(* Logix 5000 project; controller _GigaDiscovery vendor 1 type 14 code 244 rev 35.11; software revision 35.03 *) (continued)
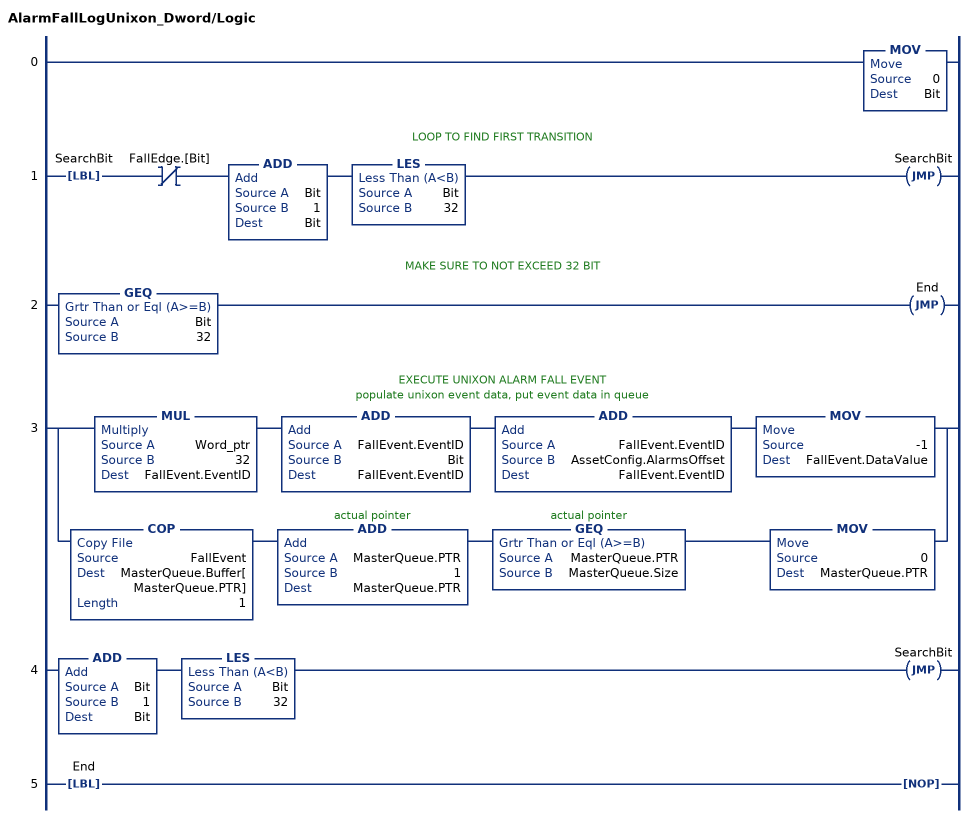
   0: MOV(0,Bit);
   // LOOP TO FIND FIRST TRANSITION
   1: LBL(SearchBit)XIO(FallEdge.[Bit])ADD(Bit,1,Bit)LES(Bit,32)JMP(SearchBit);
   // MAKE SURE TO NOT EXCEED 32 BIT
   2: GEQ(Bit,32)JMP(End);
   // EXECUTE UNIXON ALARM FALL EVENT
   // populate unixon event data, put event data in queue
   3: [MUL(Word_ptr,32,FallEvent.EventID) ADD(FallEvent.EventID,Bit,FallEvent.EventID) ADD(FallEvent.EventID,AssetConfig.AlarmsOffset,FallEvent.EventID) MOV(-1,FallEvent.DataValue) ,COP(FallEvent,MasterQueue.Buffer[MasterQueue.PTR],1) ADD(MasterQueue.PTR,1,MasterQueue.PTR) GEQ(MasterQueue.PTR,MasterQueue.Size) MOV(0,MasterQueue.PTR) ];
   4: ADD(Bit,1,Bit)LES(Bit,32)JMP(SearchBit);
   5: LBL(End)NOP();
END_ROUTINE
END_ADD_ON_INSTRUCTION

ADD_ON_INSTRUCTION AOI_DCM   (* revision 1.0 *)
VAR_INPUT
   Input_Type : BOOL; {required}   // 0 = Equivalent 1 = Complementary
   Discrepancy_Time : DINT; {required}   // (Msec)
   Channel_A : BOOL; {required}
   Channel_B : BOOL; {required}
   Channel_A_Status : BOOL; {required}
   Channel_B_Status : BOOL; {required}
   Reset_Pulse : BOOL; {required}
END_VAR
VAR_OUTPUT
   O1 : BOOL; {access Read Only, visible}
   FP : BOOL; {visible}
END_VAR
VAR
   Discrepancy_Timer : TIMER; {access None}
   Os : BOOL; {access None}
END_VAR

ROUTINE Logic   (* ladder *)
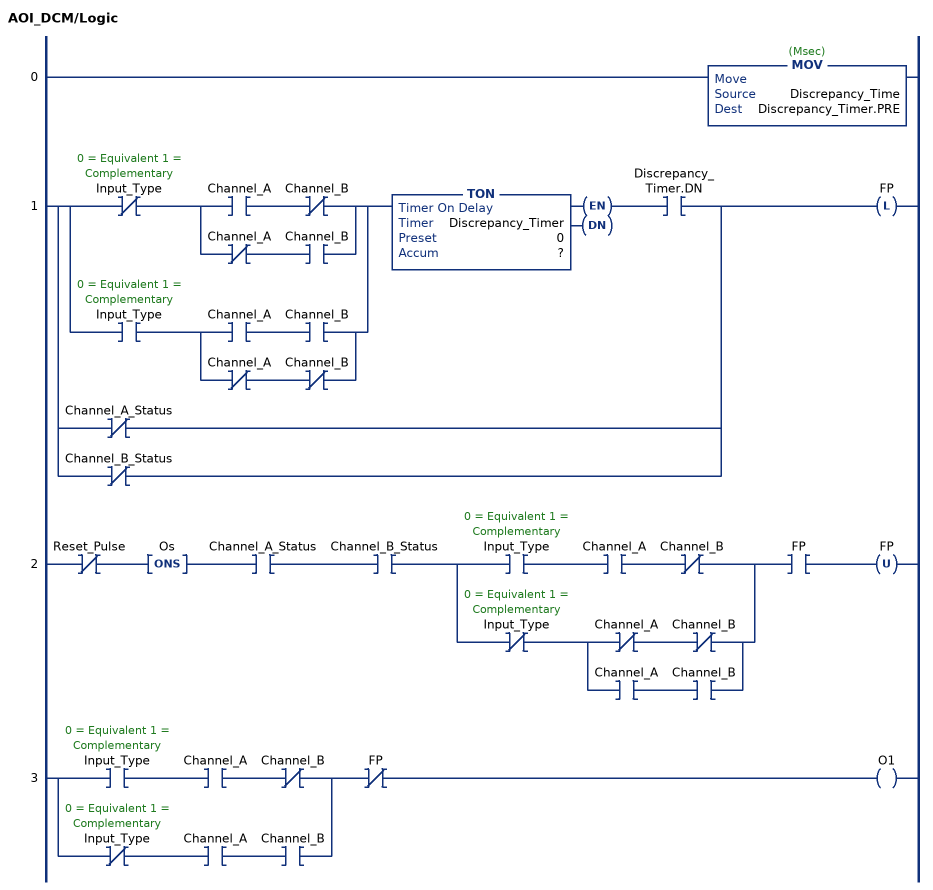
   0: MOV(Discrepancy_Time,Discrepancy_Timer.PRE);
   1: [[XIO(Input_Type) [XIC(Channel_A) XIO(Channel_B) ,XIO(Channel_A) XIC(Channel_B) ] ,XIC(Input_Type) [XIC(Channel_A) XIC(Channel_B) ,XIO(Channel_A) XIO(Channel_B) ] ] TON(Discrepancy_Timer,?,?) XIC(Discrepancy_Timer.DN) ,XIO(Channel_A_Status) ,XIO(Channel_B_Status) ]OTL(FP);
   2: XIO(Reset_Pulse)ONS(Os)XIC(Channel_A_Status)XIC(Channel_B_Status)[XIC(Input_Type) XIC(Channel_A) XIO(Channel_B) ,XIO(Input_Type) [XIO(Channel_A) XIO(Channel_B) ,XIC(Channel_A) XIC(Channel_B) ] ]XIC(FP)OTU(FP);
   3: [XIC(Input_Type) XIC(Channel_A) XIO(Channel_B) ,XIO(Input_Type) XIC(Channel_A) XIC(Channel_B) ]XIO(FP)OTE(O1);
END_ROUTINE
END_ADD_ON_INSTRUCTION

ADD_ON_INSTRUCTION EStop_AOI   (* revision 1.0, vendor Auxel *)
// Test the E-Stop Push Botton
// Revision note:
// Preliminary
// Help:
// This AOI request at the operator to check hte E-Stop function in cold mode (Ride not in start mode)
VAR_INPUT
   InEStopPbCh1 : BOOL; {access None, required}
   InEStopPbCh2 : BOOL; {required}
   InStatusCh1 : BOOL; {required}
   InStatusCh2 : BOOL; {required}
   cmdFltRst : BOOL; {required}
END_VAR
VAR_OUTPUT
   Test_Ok : BOOL; {access Read Only, visible}   // Test succefuly
   O1 : BOOL; {visible}
   FP : BOOL; {access Read Only, visible}
END_VAR
VAR
   Os : DINT; {access None}
   Sequencer : DINT; {access None}
   DCIS : DCI_STOP; {access None}
   In_Status : BOOL; {access None}
   PowerON : TIMER := (PRE := 200); {access None}
END_VAR

ROUTINE Logic   (* ladder *)
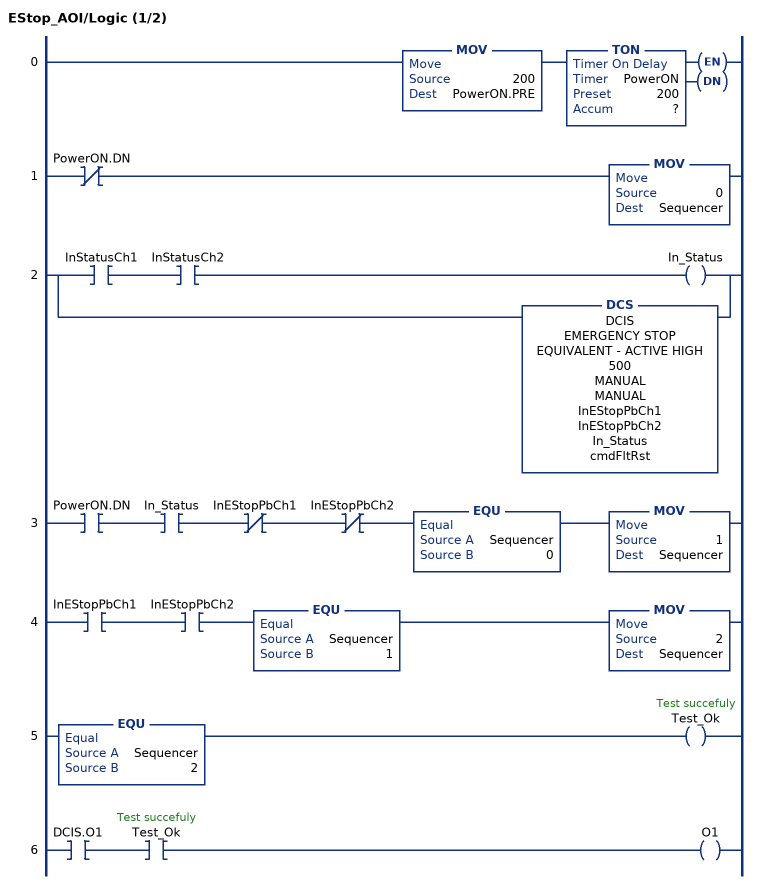
   0: MOV(200,PowerON.PRE)TON(PowerON,?,?);
   1: XIO(PowerON.DN)MOV(0,Sequencer);
   2: [XIC(InStatusCh1) XIC(InStatusCh2) OTE(In_Status) ,DCS(DCIS,EMERGENCY STOP,EQUIVALENT - ACTIVE HIGH,500,MANUAL,MANUAL,InEStopPbCh1,InEStopPbCh2,In_Status,cmdFltRst) ];
   3: XIC(PowerON.DN)XIC(In_Status)XIO(InEStopPbCh1)XIO(InEStopPbCh2)EQU(Sequencer,0)MOV(1,Sequencer);
   4: XIC(InEStopPbCh1)XIC(InEStopPbCh2)EQU(Sequencer,1)MOV(2,Sequencer);
   5: EQU(Sequencer,2)OTE(Test_Ok);
   6: XIC(DCIS.O1)XIC(Test_Ok)OTE(O1);
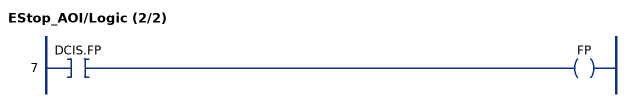
   7: XIC(DCIS.FP)OTE(FP);
END_ROUTINE
END_ADD_ON_INSTRUCTION

ADD_ON_INSTRUCTION Life_of_Machine   (* revision 1.0 *)
VAR_INPUT
   Start_Stop_Cycle_Started : BOOL; {required}
   HMI_Reset_Partial_Life_RunHH : BOOL; {required}
   HMI_Reset_Partial_Life_Cycle : BOOL; {required}
END_VAR
VAR_OUTPUT
   Life_HH : DINT; {access Read Only, visible}
   Partial_Life_HH : DINT; {access Read Only, visible}
   Working_Cycle_Number_Partial : DINT; {access Read Only, visible}
   Working_Cycle_Number_Total : DINT; {access Read Only, visible}
   Working_HH_Partial : DINT; {access Read Only, visible}
   Working_HH_Total : DINT; {access Read Only, visible}
   Working_Minutes_Partial : DINT; {access Read Only, visible}
END_VAR
VAR_INPUT
   HMI_Reset_Life_of_Machine : BOOL;
END_VAR
VAR
   Life_Hours : TIMER := (PRE := 3600000, ACC := 2467243); {access None}
   Life_HH_CTU : COUNTER; {access None}
   Partial_Life_HH_CTU : COUNTER; {access None}
   Working_Hours : TIMER := (PRE := 3600000, ACC := 2768993); {access None}
   Working_Minutes : TIMER := (PRE := 60000, ACC := 4300); {access None}
   Working_Cycle_Number_Partial_CTU : COUNTER; {access None}
   Working_Cycle_Number_Total_CTU : COUNTER; {access None}
   Working_HH_Partial_CTU : COUNTER; {access None}
   Working_HH_Total_CTU : COUNTER; {access None}
   Working_Minutes_Partial_CTU : COUNTER; {access None}
   Os : DINT; {access None}
END_VAR

ROUTINE Logic   (* ladder *)
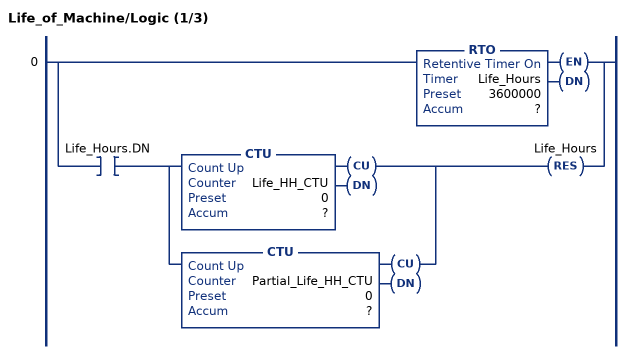
   0: [RTO(Life_Hours,?,?) ,XIC(Life_Hours.DN) [CTU(Life_HH_CTU,?,?) ,CTU(Partial_Life_HH_CTU,?,?) ] RES(Life_Hours) ];
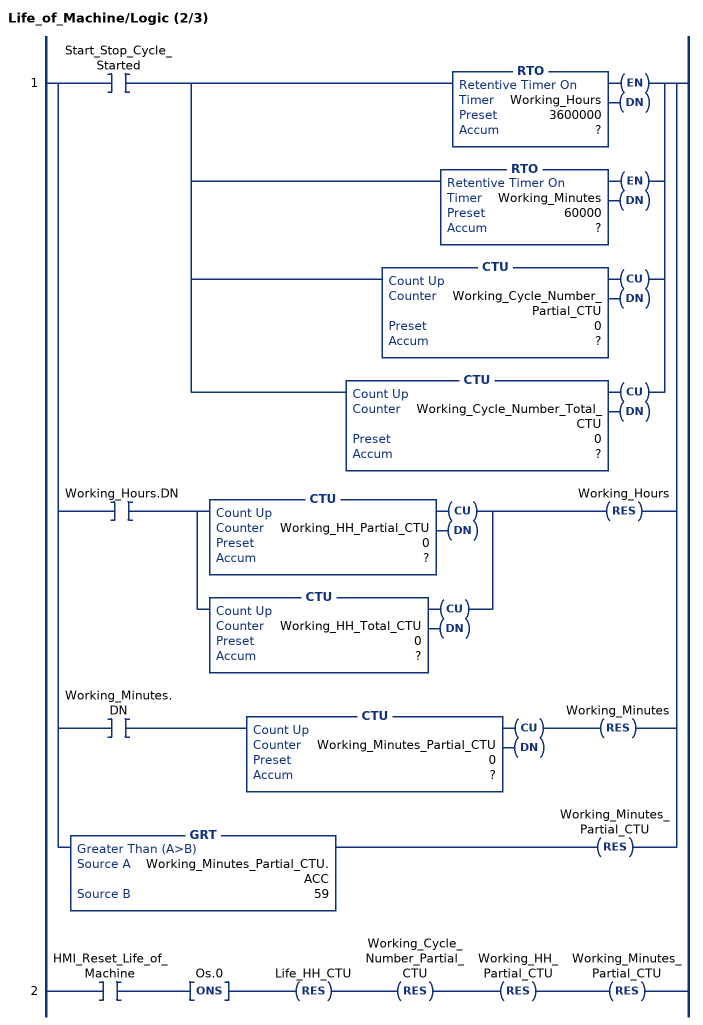
   1: [XIC(Start_Stop_Cycle_Started) [RTO(Working_Hours,?,?) ,RTO(Working_Minutes,?,?) ,[CTU(Working_Cycle_Number_Partial_CTU,?,?) ,CTU(Working_Cycle_Number_Total_CTU,?,?) ] ] ,XIC(Working_Hours.DN) [CTU(Working_HH_Partial_CTU,?,?) ,CTU(Working_HH_Total_CTU,?,?) ] RES(Working_Hours) ,XIC(Working_Minutes.DN) CTU(Working_Minutes_Partial_CTU,?,?) RES(Working_Minutes) ,GRT(Working_Minutes_Partial_CTU.ACC,59) RES(Working_Minutes_Partial_CTU) ];
   2: XIC(HMI_Reset_Life_of_Machine)ONS(Os.0)RES(Life_HH_CTU)RES(Working_Cycle_Number_Partial_CTU)RES(Working_HH_Partial_CTU)RES(Working_Minutes_Partial_CTU);
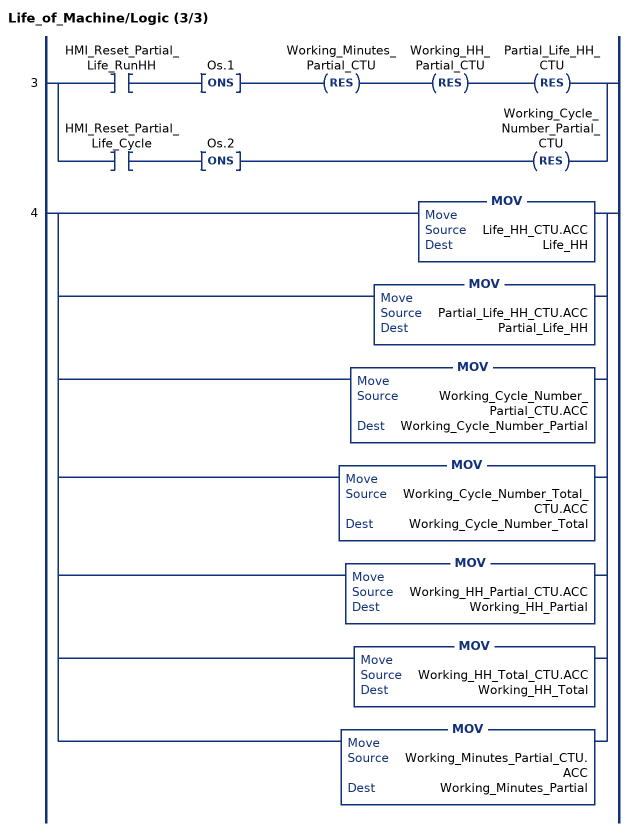
   3: [XIC(HMI_Reset_Partial_Life_RunHH) ONS(Os.1) RES(Working_Minutes_Partial_CTU) RES(Working_HH_Partial_CTU) RES(Partial_Life_HH_CTU) ,XIC(HMI_Reset_Partial_Life_Cycle) ONS(Os.2) RES(Working_Cycle_Number_Partial_CTU) ];
   4: [MOV(Life_HH_CTU.ACC,Life_HH) ,MOV(Partial_Life_HH_CTU.ACC,Partial_Life_HH) ,MOV(Working_Cycle_Number_Partial_CTU.ACC,Working_Cycle_Number_Partial) ,MOV(Working_Cycle_Number_Total_CTU.ACC,Working_Cycle_Number_Total) ,MOV(Working_HH_Partial_CTU.ACC,Working_HH_Partial) ,MOV(Working_HH_Total_CTU.ACC,Working_HH_Total) ,MOV(Working_Minutes_Partial_CTU.ACC,Working_Minutes_Partial) ];
END_ROUTINE
END_ADD_ON_INSTRUCTION

ADD_ON_INSTRUCTION Powerflex_DC_Fault   (* revision 1.0 *)
VAR_INPUT
   Fault_Code : DINT; {required}
END_VAR
VAR_IN_OUT
   Fault_Descrpition : STRING; {required}
END_VAR
VAR
   Fault_Descrpition_4 : STRING := 'AC Undervoltage'; {access None}
   Fault_Descrpition_5 : STRING := 'Arm Overvoltage'; {access None}
   Fault_Descrpition_2 : STRING := 'Auxiliary Input'; {access None}
   Fault_Descrpition_64 : STRING := 'Drive Overload'; {access None}
   Fault_Descrpition_132 : STRING := 'Dsp Error'; {access None}
   Fault_Descrpition_100 : STRING := '100'; {access None}
   Fault_Descrpition_32 : STRING; {access None}
   Fault_Descrpition_6 : STRING := 'Fld Current Loss'; {access None}
   Fault_Descrpition_95 : STRING := 'Fwd End Limit'; {access None}
   Fault_Descrpition_97 : STRING := 'Fwd Over Travel'; {access None}
   Fault_Descrpition_130 : STRING := 'Hardware Fault'; {access None}
   Fault_Descrpition_131 : STRING := 'Interrupt Error'; {access None}
   Fault_Descrpition_37 : STRING := 'Inverting Fault'; {access None}
   Fault_Descrpition_10 : STRING := 'Main Contactor'; {access None}
   Fault_Descrpition_7 : STRING := 'Motor Overload'; {access None}
   Fault_Descrpition_16 : STRING := 'Motor Over Temp'; {access None}
   Fault_Descrpition_90 : STRING := 'Open SCR'; {access None}
   Fault_Descrpition_13 : STRING := 'Overcurrent'; {access None}
   Fault_Descrpition_25 : STRING := 'Overspeed'; {access None}
   Fault_Descrpition_48 : STRING := 'Params Defaulted'; {access None}
   Fault_Descrpition_71 : STRING := 'Pommunication card fault Port 1'; {access None}
   Fault_Descrpition_81 : STRING := 'DPI port 1 stopped communicating'; {access None}
   Fault_Descrpition_93 : STRING := 'Resolver Error'; {access None}
   Fault_Descrpition_96 : STRING := 'Rev End Limit'; {access None}
   Fault_Descrpition_98 : STRING := 'Rev Over Travel'; {access None}
   Fault_Descrpition_89 : STRING := 'Shorted SCR'; {access None}
   Fault_Descrpition_91 : STRING := 'Spd Fdbk Loss'; {access None}
   Fault_Descrpition_62 : STRING := 'STune Aborted'; {access None}
   Fault_Descrpition_59 : STRING := 'STune CurLimit'; {access None}
   Fault_Descrpition_60 : STRING := 'STune FrictionLo'; {access None}
   Fault_Descrpition_58 : STRING := 'STune LoadHi'; {access None}
   Fault_Descrpition_56 : STRING := 'STune Overspeed'; {access None}
   Fault_Descrpition_57 : STRING := 'STune Stalled'; {access None}
   Fault_Descrpition_61 : STRING := 'STune Timeout'; {access None}
   Fault_Descrpition_70 : STRING := 'Sustained Curr'; {access None}
   Fault_Descrpition_94 : STRING := 'TorqPrv Spd Band'; {access None}
   Fault_Descrpition_99 : STRING := 'Travel Lim Cflct'; {access None}
   Fault_Descrpition_92 : STRING := 'Encoder Error'; {access None}
   Fault_Descrpition_8 : STRING := 'Heatsink OvrTemp'; {access None}
   Fault_Descrpition_82 : STRING := 'DPI port 2 stopped communicating'; {access None}
   Fault_Descrpition_83 : STRING := 'DPI port 3 stopped communicating'; {access None}
   Fault_Descrpition_84 : STRING := 'DPI port 4 stopped communicating'; {access None}
   Fault_Descrpition_85 : STRING := 'DPI port 5 stopped communicating'; {access None}
   Fault_Descrpition_72 : STRING := 'Pommunication card fault Port 2'; {access None}
   Fault_Descrpition_73 : STRING := 'Pommunication card fault Port 3'; {access None}
   Fault_Descrpition_74 : STRING := 'Pommunication card fault Port 4'; {access None}
   Fault_Descrpition_75 : STRING := 'Pommunication card fault Port 5'; {access None}
   Fault_Descrpition_3 : STRING := 'Power Failure'; {access None}
END_VAR

ROUTINE Logic   (* structured text *)
   DELETE(Fault_Descrpition,32,1,Fault_Descrpition );
   case Fault_Code of
   	4:		INSERT(Fault_Descrpition,Fault_Descrpition_4 , 1,Fault_Descrpition );
   	5:		INSERT(Fault_Descrpition,Fault_Descrpition_5 , 1,Fault_Descrpition );
   	2:		INSERT(Fault_Descrpition,Fault_Descrpition_2 , 1,Fault_Descrpition );
   	64:		INSERT(Fault_Descrpition,Fault_Descrpition_64 , 1,Fault_Descrpition );
   	132:	INSERT(Fault_Descrpition,Fault_Descrpition_132 , 1,Fault_Descrpition );
   	100:	INSERT(Fault_Descrpition,Fault_Descrpition_100 , 1,Fault_Descrpition );
   	92:		INSERT(Fault_Descrpition,Fault_Descrpition_32 , 1,Fault_Descrpition );
   	6:		INSERT(Fault_Descrpition,Fault_Descrpition_6 , 1,Fault_Descrpition );
   	95:		INSERT(Fault_Descrpition,Fault_Descrpition_95 , 1,Fault_Descrpition );
   	97:		INSERT(Fault_Descrpition,Fault_Descrpition_97 , 1,Fault_Descrpition );
   	8:		INSERT(Fault_Descrpition,Fault_Descrpition_8 , 1,Fault_Descrpition );
   	130:	INSERT(Fault_Descrpition,Fault_Descrpition_130 , 1,Fault_Descrpition );
   	131:	INSERT(Fault_Descrpition,Fault_Descrpition_131 , 1,Fault_Descrpition );
   	37:		INSERT(Fault_Descrpition,Fault_Descrpition_37 , 1,Fault_Descrpition );
   	10:		INSERT(Fault_Descrpition,Fault_Descrpition_10 , 1,Fault_Descrpition );
   	7:		INSERT(Fault_Descrpition,Fault_Descrpition_7 , 1,Fault_Descrpition );
   	16:		INSERT(Fault_Descrpition,Fault_Descrpition_16 , 1,Fault_Descrpition );
   	90:		INSERT(Fault_Descrpition,Fault_Descrpition_90 , 1,Fault_Descrpition );
   	13:		INSERT(Fault_Descrpition,Fault_Descrpition_13 , 1,Fault_Descrpition );
   	25:		INSERT(Fault_Descrpition,Fault_Descrpition_25 , 1,Fault_Descrpition );
   	48:		INSERT(Fault_Descrpition,Fault_Descrpition_48 , 1,Fault_Descrpition );
   	71:		INSERT(Fault_Descrpition,Fault_Descrpition_71 , 1,Fault_Descrpition );
   	72:		INSERT(Fault_Descrpition,Fault_Descrpition_72 , 1,Fault_Descrpition );
   	73:		INSERT(Fault_Descrpition,Fault_Descrpition_73 , 1,Fault_Descrpition );
   	74:		INSERT(Fault_Descrpition,Fault_Descrpition_74 , 1,Fault_Descrpition );
   	75:		INSERT(Fault_Descrpition,Fault_Descrpition_75 , 1,Fault_Descrpition );
   	81:		INSERT(Fault_Descrpition,Fault_Descrpition_81 , 1,Fault_Descrpition );
   	82:		INSERT(Fault_Descrpition,Fault_Descrpition_82 , 1,Fault_Descrpition );
   	83:		INSERT(Fault_Descrpition,Fault_Descrpition_83 , 1,Fault_Descrpition );
   	84:		INSERT(Fault_Descrpition,Fault_Descrpition_84 , 1,Fault_Descrpition );
   	85:		INSERT(Fault_Descrpition,Fault_Descrpition_85 , 1,Fault_Descrpition );
   	3:		INSERT(Fault_Descrpition,Fault_Descrpition_3 , 1,Fault_Descrpition );
   	93:		INSERT(Fault_Descrpition,Fault_Descrpition_93 , 1,Fault_Descrpition );
   	96:		INSERT(Fault_Descrpition,Fault_Descrpition_94 , 1,Fault_Descrpition );
   	98:		INSERT(Fault_Descrpition,Fault_Descrpition_98 , 1,Fault_Descrpition );
   	89:		INSERT(Fault_Descrpition,Fault_Descrpition_89 , 1,Fault_Descrpition );
   	91:		INSERT(Fault_Descrpition,Fault_Descrpition_91 , 1,Fault_Descrpition );
   	92:		INSERT(Fault_Descrpition,Fault_Descrpition_92 , 1,Fault_Descrpition );
   	62:		INSERT(Fault_Descrpition,Fault_Descrpition_62 , 1,Fault_Descrpition );
   	59:		INSERT(Fault_Descrpition,Fault_Descrpition_59 , 1,Fault_Descrpition );
   	60:		INSERT(Fault_Descrpition,Fault_Descrpition_60 , 1,Fault_Descrpition );
   	58:		INSERT(Fault_Descrpition,Fault_Descrpition_58 , 1,Fault_Descrpition );
   	56:		INSERT(Fault_Descrpition,Fault_Descrpition_56 , 1,Fault_Descrpition );
   	57:		INSERT(Fault_Descrpition,Fault_Descrpition_57 , 1,Fault_Descrpition );
   	61:		INSERT(Fault_Descrpition,Fault_Descrpition_61 , 1,Fault_Descrpition );
   	70:		INSERT(Fault_Descrpition,Fault_Descrpition_70 , 1,Fault_Descrpition );
   	94:		INSERT(Fault_Descrpition,Fault_Descrpition_94 , 1,Fault_Descrpition );
   	99:		INSERT(Fault_Descrpition,Fault_Descrpition_99 , 1,Fault_Descrpition );
   end_case;
   
   
END_ROUTINE
END_ADD_ON_INSTRUCTION

ADD_ON_INSTRUCTION Sel_3_Pos_2_Input   (* revision 1.0 *)
VAR_INPUT
   Ch_1 : BOOL; {required}
   Ch_2 : BOOL; {required}
   Status_Ch_1 : BOOL; {required}
   Status_Ch_2 : BOOL; {required}
END_VAR
VAR_OUTPUT
   Left : BOOL; {access None, visible}
   Center : BOOL; {access None, visible}
   Right : BOOL; {access None, visible}
   Fault : BOOL; {access None, visible}
END_VAR
VAR_INPUT
   Alarm_Reset : BOOL; {required}
END_VAR
VAR
   Channels_Status : BOOL; {access None}
   Timer : TIMER := (PRE := 2500); {access None}
END_VAR

ROUTINE Logic   (* ladder *)
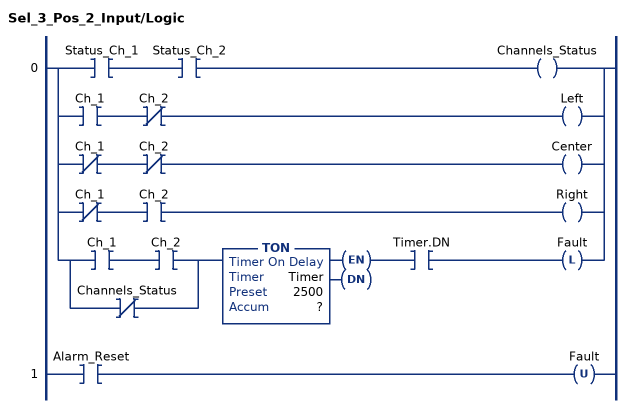
   0: [XIC(Status_Ch_1) XIC(Status_Ch_2) OTE(Channels_Status) ,XIC(Ch_1) XIO(Ch_2) OTE(Left) ,XIO(Ch_1) XIO(Ch_2) OTE(Center) ,XIO(Ch_1) XIC(Ch_2) OTE(Right) ,[XIC(Ch_1) XIC(Ch_2) ,XIO(Channels_Status) ] TON(Timer,?,?) XIC(Timer.DN) OTL(Fault) ];
   1: XIC(Alarm_Reset)OTU(Fault);
END_ROUTINE
END_ADD_ON_INSTRUCTION

ADD_ON_INSTRUCTION Sel_3_Pos_3_Input   (* revision 1.0 *)
VAR_INPUT
   Ch_1 : BOOL; {required}
   Ch_2 : BOOL; {required}
   Ch_3 : BOOL; {required}
   Status_Ch_1 : BOOL; {required}
   Status_Ch_2 : BOOL; {required}
   Status_Ch_3 : BOOL; {required}
END_VAR
VAR_OUTPUT
   Left : BOOL; {access None, visible}
   Center : BOOL; {access None, visible}
   Right : BOOL; {access None, visible}
   Fault : BOOL; {access None, visible}
END_VAR
VAR_INPUT
   Alarm_Reset : BOOL; {required}
END_VAR
VAR
   Channels_Status : BOOL; {access None}
   Timer : TIMER := (PRE := 2500); {access None}
END_VAR

ROUTINE Logic   (* ladder *)
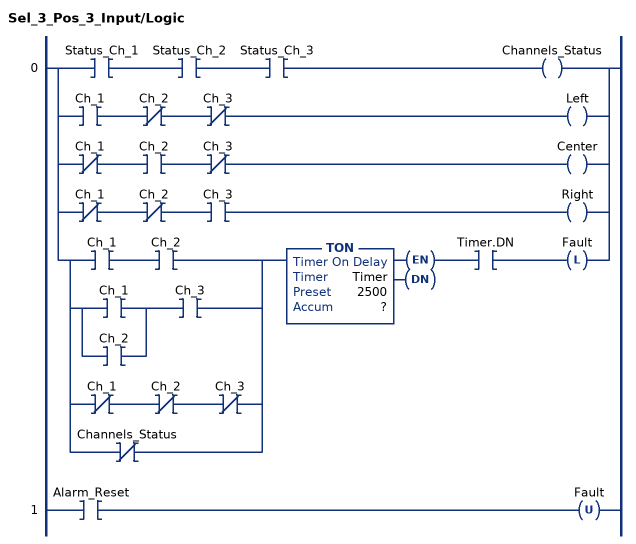
   0: [XIC(Status_Ch_1) XIC(Status_Ch_2) XIC(Status_Ch_3) OTE(Channels_Status) ,XIC(Ch_1) XIO(Ch_2) XIO(Ch_3) OTE(Left) ,XIO(Ch_1) XIC(Ch_2) XIO(Ch_3) OTE(Center) ,XIO(Ch_1) XIO(Ch_2) XIC(Ch_3) OTE(Right) ,[XIC(Ch_1) XIC(Ch_2) ,[XIC(Ch_1) ,XIC(Ch_2) ] XIC(Ch_3) ,XIO(Ch_1) XIO(Ch_2) XIO(Ch_3) ,XIO(Channels_Status) ] TON(Timer,?,?) XIC(Timer.DN) OTL(Fault) ];
   1: XIC(Alarm_Reset)OTU(Fault);
END_ROUTINE
END_ADD_ON_INSTRUCTION

ADD_ON_INSTRUCTION Sequencer_AOI   (* revision 1.0 *)
VAR_IN_OUT
   DataInOut : Sequencer; {required}
END_VAR
VAR
   Timer_start_OFF_Delay : TIMER := (PRE := 200); {access None}
END_VAR

ROUTINE Logic   (* ladder *)
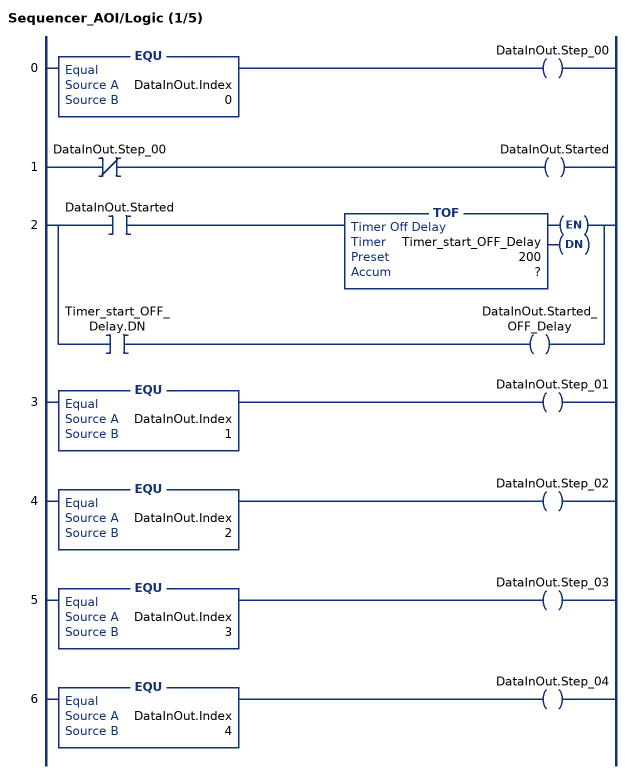
   0: EQU(DataInOut.Index,0)OTE(DataInOut.Step_00);
   1: XIO(DataInOut.Step_00)OTE(DataInOut.Started);
   2: [XIC(DataInOut.Started) TOF(Timer_start_OFF_Delay,?,?) ,XIC(Timer_start_OFF_Delay.DN) OTE(DataInOut.Started_OFF_Delay) ];
   3: EQU(DataInOut.Index,1)OTE(DataInOut.Step_01);
   4: EQU(DataInOut.Index,2)OTE(DataInOut.Step_02);
   5: EQU(DataInOut.Index,3)OTE(DataInOut.Step_03);
   6: EQU(DataInOut.Index,4)OTE(DataInOut.Step_04);
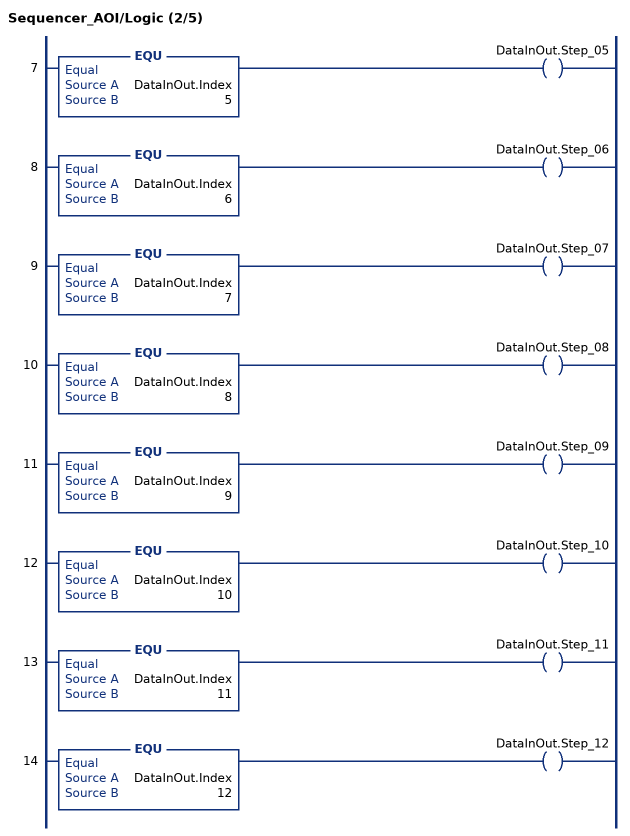
   7: EQU(DataInOut.Index,5)OTE(DataInOut.Step_05);
   8: EQU(DataInOut.Index,6)OTE(DataInOut.Step_06);
   9: EQU(DataInOut.Index,7)OTE(DataInOut.Step_07);
   10: EQU(DataInOut.Index,8)OTE(DataInOut.Step_08);
   11: EQU(DataInOut.Index,9)OTE(DataInOut.Step_09);
   12: EQU(DataInOut.Index,10)OTE(DataInOut.Step_10);
   13: EQU(DataInOut.Index,11)OTE(DataInOut.Step_11);
   14: EQU(DataInOut.Index,12)OTE(DataInOut.Step_12);
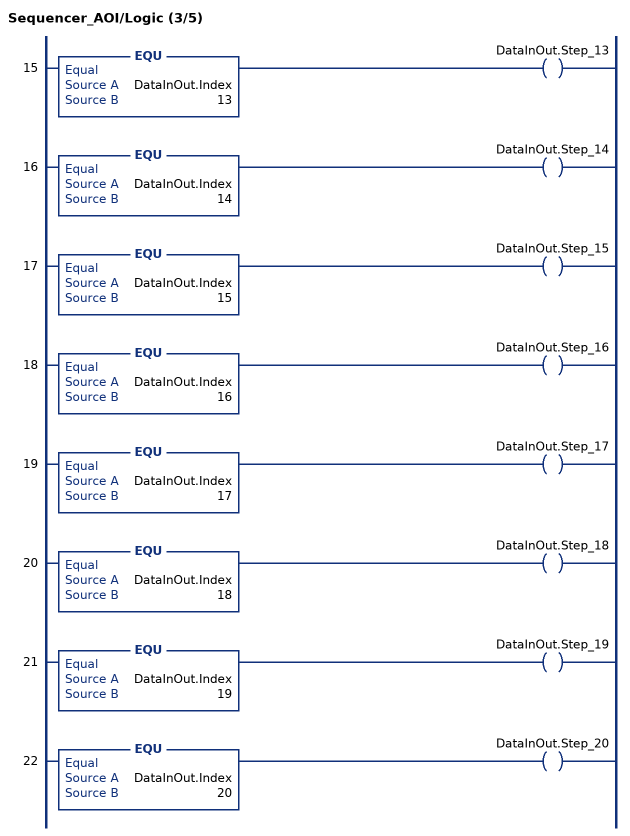
   15: EQU(DataInOut.Index,13)OTE(DataInOut.Step_13);
   16: EQU(DataInOut.Index,14)OTE(DataInOut.Step_14);
   17: EQU(DataInOut.Index,15)OTE(DataInOut.Step_15);
   18: EQU(DataInOut.Index,16)OTE(DataInOut.Step_16);
   19: EQU(DataInOut.Index,17)OTE(DataInOut.Step_17);
   20: EQU(DataInOut.Index,18)OTE(DataInOut.Step_18);
   21: EQU(DataInOut.Index,19)OTE(DataInOut.Step_19);
   22: EQU(DataInOut.Index,20)OTE(DataInOut.Step_20);
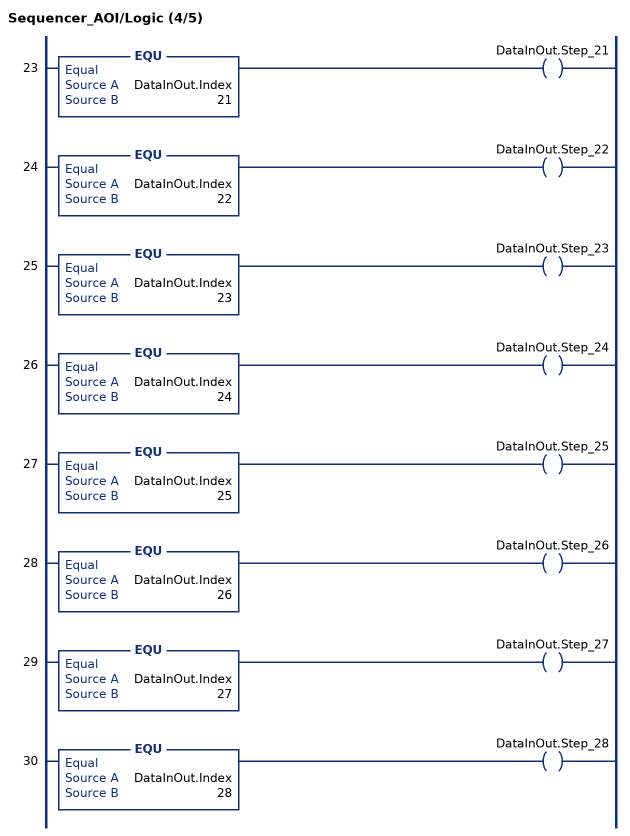
   23: EQU(DataInOut.Index,21)OTE(DataInOut.Step_21);
   24: EQU(DataInOut.Index,22)OTE(DataInOut.Step_22);
   25: EQU(DataInOut.Index,23)OTE(DataInOut.Step_23);
   26: EQU(DataInOut.Index,24)OTE(DataInOut.Step_24);
   27: EQU(DataInOut.Index,25)OTE(DataInOut.Step_25);
   28: EQU(DataInOut.Index,26)OTE(DataInOut.Step_26);
   29: EQU(DataInOut.Index,27)OTE(DataInOut.Step_27);
   30: EQU(DataInOut.Index,28)OTE(DataInOut.Step_28);
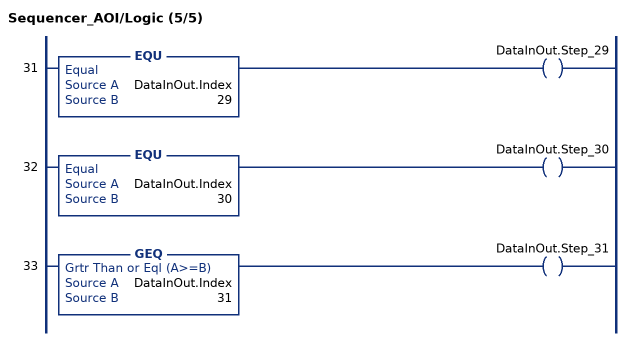
   31: EQU(DataInOut.Index,29)OTE(DataInOut.Step_29);
   32: EQU(DataInOut.Index,30)OTE(DataInOut.Step_30);
   33: GEQ(DataInOut.Index,31)OTE(DataInOut.Step_31);
END_ROUTINE
END_ADD_ON_INSTRUCTION

ADD_ON_INSTRUCTION Sequencer_AOI_Std   (* revision 1.0 *)
VAR_IN_OUT
   DataInOut : Sequencer; {required}
END_VAR
VAR
   Timer_start_OFF_Delay : TIMER := (PRE := 200); {access None}
END_VAR

ROUTINE Logic   (* ladder *)
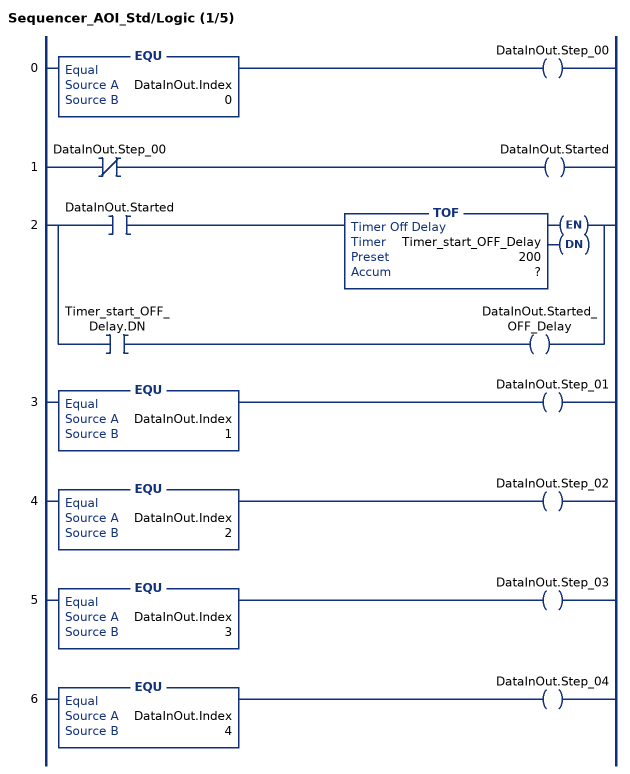
   0: EQU(DataInOut.Index,0)OTE(DataInOut.Step_00);
   1: XIO(DataInOut.Step_00)OTE(DataInOut.Started);
   2: [XIC(DataInOut.Started) TOF(Timer_start_OFF_Delay,?,?) ,XIC(Timer_start_OFF_Delay.DN) OTE(DataInOut.Started_OFF_Delay) ];
   3: EQU(DataInOut.Index,1)OTE(DataInOut.Step_01);
   4: EQU(DataInOut.Index,2)OTE(DataInOut.Step_02);
   5: EQU(DataInOut.Index,3)OTE(DataInOut.Step_03);
   6: EQU(DataInOut.Index,4)OTE(DataInOut.Step_04);
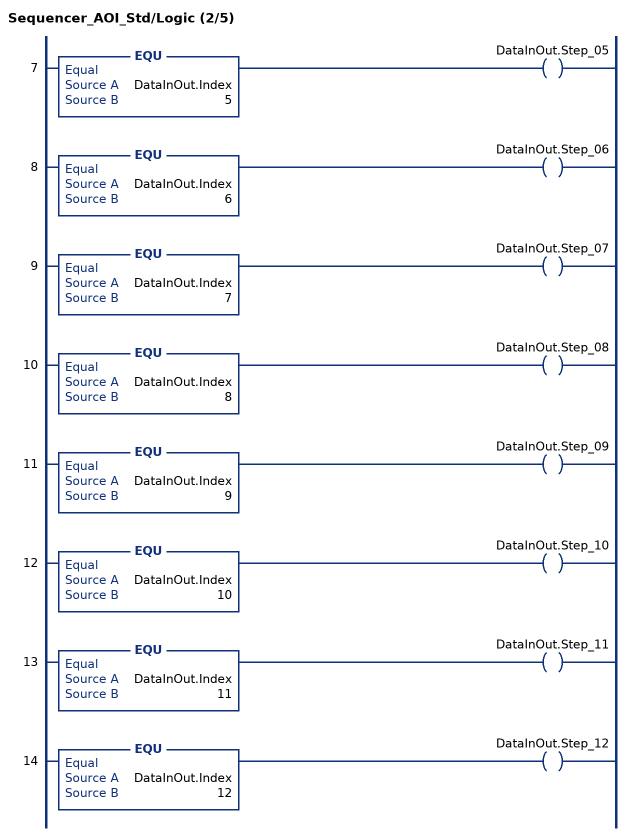
   7: EQU(DataInOut.Index,5)OTE(DataInOut.Step_05);
   8: EQU(DataInOut.Index,6)OTE(DataInOut.Step_06);
   9: EQU(DataInOut.Index,7)OTE(DataInOut.Step_07);
   10: EQU(DataInOut.Index,8)OTE(DataInOut.Step_08);
   11: EQU(DataInOut.Index,9)OTE(DataInOut.Step_09);
   12: EQU(DataInOut.Index,10)OTE(DataInOut.Step_10);
   13: EQU(DataInOut.Index,11)OTE(DataInOut.Step_11);
   14: EQU(DataInOut.Index,12)OTE(DataInOut.Step_12);
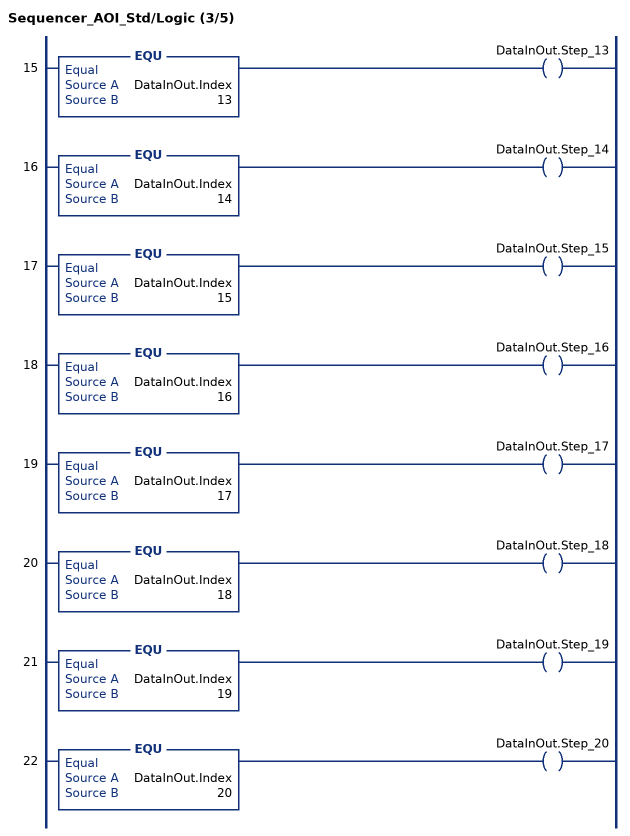
   15: EQU(DataInOut.Index,13)OTE(DataInOut.Step_13);
   16: EQU(DataInOut.Index,14)OTE(DataInOut.Step_14);
   17: EQU(DataInOut.Index,15)OTE(DataInOut.Step_15);
   18: EQU(DataInOut.Index,16)OTE(DataInOut.Step_16);
   19: EQU(DataInOut.Index,17)OTE(DataInOut.Step_17);
   20: EQU(DataInOut.Index,18)OTE(DataInOut.Step_18);
   21: EQU(DataInOut.Index,19)OTE(DataInOut.Step_19);
   22: EQU(DataInOut.Index,20)OTE(DataInOut.Step_20);
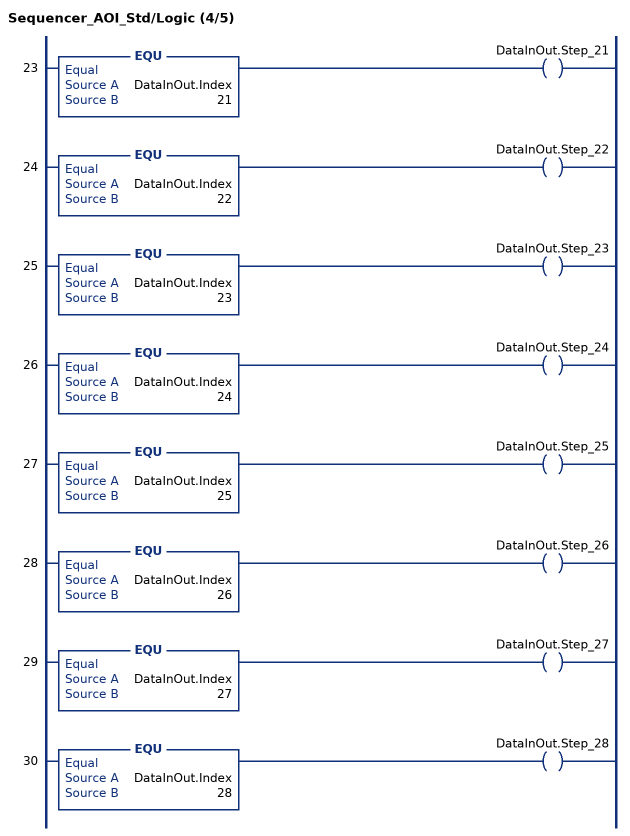
   23: EQU(DataInOut.Index,21)OTE(DataInOut.Step_21);
   24: EQU(DataInOut.Index,22)OTE(DataInOut.Step_22);
   25: EQU(DataInOut.Index,23)OTE(DataInOut.Step_23);
   26: EQU(DataInOut.Index,24)OTE(DataInOut.Step_24);
   27: EQU(DataInOut.Index,25)OTE(DataInOut.Step_25);
   28: EQU(DataInOut.Index,26)OTE(DataInOut.Step_26);
   29: EQU(DataInOut.Index,27)OTE(DataInOut.Step_27);
   30: EQU(DataInOut.Index,28)OTE(DataInOut.Step_28);
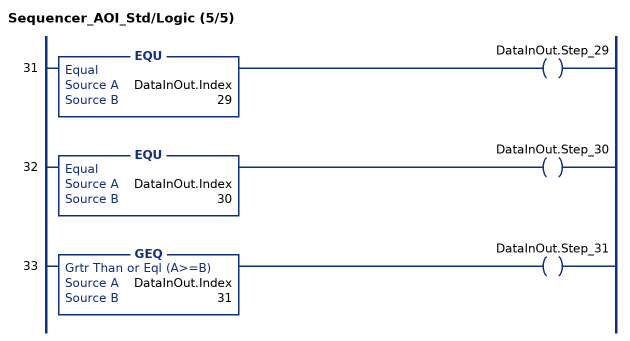
   31: EQU(DataInOut.Index,29)OTE(DataInOut.Step_29);
   32: EQU(DataInOut.Index,30)OTE(DataInOut.Step_30);
   33: GEQ(DataInOut.Index,31)OTE(DataInOut.Step_31);
END_ROUTINE
END_ADD_ON_INSTRUCTION
